screen "Manual.General" 800x480, template "TemplateWithClockAndBackBtnForManual"
   on GenerateScreen: SetBit("Maintenance")
   on ClearScreen: ResetBit("Maintenance")
   GraphicIOField "PlotLight_Round_G" at 224,264 size 24x24; PictureOff "PilotLight_Round_G_Off_256c"; PictureOn "PilotLight_Round_G_On_256c"
      ProcessValue <- "Prezenta aer"
   TextField "Text field_1" at 8,266 size 90x20; Text 'Prezenta aer'
   GraphicIOField "PlotLight_Round_G_1" at 224,48 size 24x24; PictureOn "PilotLight_Round_G_On_256c"; PictureOff "PilotLight_Round_G_Off_256c"
      ProcessValue <- "Aliniere palet"
   TextField "Text field_2" at 8,50 size 91x20; Text 'Aliniere palet'
   GraphicIOField "PlotLight_Round_G_2" at 224,72 size 24x24; PictureOff "PilotLight_Round_G_Off_256c"; PictureOn "PilotLight_Round_G_On_256c"
      ProcessValue <- "Centror extins"
   TextField "Text field_3" at 8,74 size 98x20; Text 'Centror extins'
   GraphicIOField "PlotLight_Round_G_3" at 224,96 size 24x24; PictureOff "PilotLight_Round_G_Off_256c"; PictureOn "PilotLight_Round_G_On_256c"
      ProcessValue <- "Centror retras"
   TextField "Text field_4" at 8,98 size 100x20; Text 'Centror retras'
   GraphicIOField "PlotLight_Round_G_4" at 224,120 size 24x24; PictureOff "PilotLight_Round_G_Off_256c"; PictureOn "PilotLight_Round_G_On_256c"
      ProcessValue <- "Detectie 1 aliniament palet"
   TextField "Text field_5" at 8,122 size 179x20; Text 'Detectie 1 aliniament palet'
   GraphicIOField "PlotLight_Round_G_5" at 224,144 size 24x24; PictureOff "PilotLight_Round_G_Off_256c"; PictureOn "PilotLight_Round_G_On_256c"
      ProcessValue <- "Detectie 2 aliniament palet"
   TextField "Text field_6" at 8,146 size 179x20; Text 'Detectie 2 aliniament palet'
   GraphicIOField "PlotLight_Round_G_6" at 224,168 size 24x24; PictureOff "PilotLight_Round_G_Off_256c"; PictureOn "PilotLight_Round_G_On_256c"
      ProcessValue <- "Detectie palet"
   TextField "Text field_7" at 8,170 size 97x20; Text 'Detectie palet'
   GraphicIOField "PlotLight_Round_G_7" at 224,192 size 24x24; PictureOn "PilotLight_Round_G_On_256c"; PictureOff "PilotLight_Round_G_Off_256c"
      ProcessValue <- "Feed palet"
   TextField "Text field_8" at 8,194 size 72x20; Text 'Feed palet'
   GraphicIOField "PlotLight_Round_G_8" at 224,216 size 24x24; PictureOn "PilotLight_Round_G_On_256c"; PictureOff "PilotLight_Round_G_Off_256c"
      ProcessValue <- "Inaltime maxima"
   TextField "Text field_9" at 8,218 size 109x20; Text 'Inaltime maxima'
   GraphicIOField "PlotLight_Round_G_9" at 224,240 size 24x24; PictureOn "PilotLight_Round_G_On_256c"; PictureOff "PilotLight_Round_G_Off_256c"
      ProcessValue <- "Masurare lungime"
   TextField "Text field_10" at 8,242 size 120x20; Text 'Masurare lungime'
   GraphicIOField "PlotLight_Round_G_10" at 224,288 size 24x24; PictureOn "PilotLight_Round_G_On_256c"; PictureOff "PilotLight_Round_G_Off_256c"
      ProcessValue <- "Prezenta palet iesire"
   TextField "Text field_11" at 8,290 size 140x20; Text 'Prezenta palet iesire'
   GraphicIOField "PlotLight_Round_G_11" at 224,312 size 24x24; PictureOn "PilotLight_Round_G_On_256c"; PictureOff "PilotLight_Round_G_Off_256c"
      ProcessValue <- "Prezenta palet_capat_conveyor"
   TextField "Text field_12" at 8,314 size 215x20; Text 'Prezenta palet_capat_conveyor'
   GraphicIOField "PlotLight_Round_G_12" at 224,336 size 24x24; PictureOn "PilotLight_Round_G_On_256c"; PictureOff "PilotLight_Round_G_Off_256c"
      ProcessValue <- "Prezenta palet_centror"
   TextField "Text field_13" at 8,338 size 158x20; Text 'Prezenta palet_centror'
   GraphicIOField "PlotLight_Round_G_13" at 224,360 size 24x24; PictureOn "PilotLight_Round_G_On_256c"; PictureOff "PilotLight_Round_G_Off_256c"
      ProcessValue <- "Prezenta palet_dreapta"
   TextField "Text field_14" at 8,362 size 161x20; Text 'Prezenta palet_dreapta'
   GraphicIOField "PlotLight_Round_G_14" at 504,264 size 24x24; PictureOn "PilotLight_Round_G_On_256c"; PictureOff "PilotLight_Round_G_Off_256c"
      ProcessValue <- "Protectie cuplata Post reparatii minore"
   TextField "Text field_15" at 264,266 size 230x20; Text 'Prot. cuplata Post reparatii minore'
   GraphicIOField "PlotLight_Round_G_15" at 504,48 size 24x24; PictureOff "PilotLight_Round_G_Off_256c"; PictureOn "PilotLight_Round_G_On_256c"
      ProcessValue <- "Prezenta palet_stanga"
   TextField "Text field_16" at 264,50 size 154x20; Text 'Prezenta palet_stanga'
   GraphicIOField "PlotLight_Round_G_16" at 504,72 size 24x24; PictureOn "PilotLight_Round_G_On_256c"; PictureOff "PilotLight_Round_G_Off_256c"
      ProcessValue <- "Prezenta stiva"
   TextField "Text field_17" at 264,74 size 100x20; Text 'Prezenta stiva'
   GraphicIOField "PlotLight_Round_G_17" at 504,96 size 24x24; PictureOn "PilotLight_Round_G_On_256c"; PictureOff "PilotLight_Round_G_Off_256c"
      ProcessValue <- "Prezenta_stiva"
   TextField "Text field_18" at 264,98 size 104x20; Text 'Prezenta_stiva'
   GraphicIOField "PlotLight_Round_G_18" at 504,120 size 24x24; PictureOn "PilotLight_Round_G_On_256c"; PictureOff "PilotLight_Round_G_Off_256c"
      ProcessValue <- "Protectie cuplata Circular masa fixa"
   TextField "Text field_19" at 264,122 size 235x20; Text 'Protectie cuplata Circular masa fixa'
   GraphicIOField "PlotLight_Round_G_19" at 504,144 size 24x24; PictureOn "PilotLight_Round_G_On_256c"; PictureOff "PilotLight_Round_G_Off_256c"
      ProcessValue <- "Protectie cuplata HMI"
   TextField "Text field_20" at 264,146 size 146x20; Text 'Protectie cuplata HMI'
   GraphicIOField "PlotLight_Round_G_20" at 504,168 size 24x24; PictureOn "PilotLight_Round_G_On_256c"; PictureOff "PilotLight_Round_G_Off_256c"
      ProcessValue <- "Protectie cuplata Iluminat"
   TextField "Text field_21" at 264,170 size 173x20; Text 'Protectie cuplata Iluminat'
   GraphicIOField "PlotLight_Round_G_21" at 504,192 size 24x24; PictureOff "PilotLight_Round_G_Off_256c"; PictureOn "PilotLight_Round_G_On_256c"
      ProcessValue <- "Protectie cuplata Masina demontare paleti dreapta"
   TextField "Text field_22" at 264,194 size 241x20; Text 'Prot. cuplata Mas. dem. pal. dreapta'
   GraphicIOField "PlotLight_Round_G_22" at 504,216 size 24x24; PictureOff "PilotLight_Round_G_Off_256c"; PictureOn "PilotLight_Round_G_On_256c"
      ProcessValue <- "Protectie cuplata Masina demontare paleti stanga"
   TextField "Text field_23" at 264,218 size 234x20; Text 'Prot. cuplata Mas. dem. pal. stanga'
   GraphicIOField "PlotLight_Round_G_23" at 504,240 size 24x24; PictureOff "PilotLight_Round_G_Off_256c"; PictureOn "PilotLight_Round_G_On_256c"
      ProcessValue <- "Protectie cuplata Post reparatie stanga+dreapta"
   TextField "Text field_24" at 264,242 size 218x20; Text 'Prot. cuplata Post rep. stg.+drp.'
   GraphicIOField "PlotLight_Round_G_24" at 504,288 size 24x24; PictureOff "PilotLight_Round_G_Off_256c"; PictureOn "PilotLight_Round_G_On_256c"
      ProcessValue <- "Protectie cuplata TELE"
   TextField "Text field_25" at 264,290 size 149x20; Text 'Protectie cuplata TELE'
   GraphicIOField "PlotLight_Round_G_25" at 504,312 size 24x24; PictureOff "PilotLight_Round_G_Off_256c"; PictureOn "PilotLight_Round_G_On_256c"
      ProcessValue <- "Prezenta palet_capat_conveyor"
   TextField "Text field_26" at 264,314 size 215x20; Text 'Prezenta palet_capat_conveyor'
   GraphicIOField "PlotLight_Round_G_26" at 504,336 size 24x24; PictureOff "PilotLight_Round_G_Off_256c"; PictureOn "PilotLight_Round_G_On_256c"
      ProcessValue <- "Prezenta palet_centror"
   TextField "Text field_27" at 264,338 size 158x20; Text 'Prezenta palet_centror'
   GraphicIOField "PlotLight_Round_G_27" at 504,360 size 24x24; PictureOff "PilotLight_Round_G_Off_256c"; PictureOn "PilotLight_Round_G_On_256c"
      ProcessValue <- "Prezenta palet_dreapta"
   TextField "Text field_28" at 264,362 size 161x20; Text 'Prezenta palet_dreapta'
   GraphicIOField "PlotLight_Round_G_28" at 760,48 size 24x24; PictureOn "PilotLight_Round_G_On_256c"; PictureOff "PilotLight_Round_G_Off_256c"
      ProcessValue <- "Senzor 1 prezenta stiva"
   TextField "Text field_29" at 544,50 size 161x20; Text 'Senzor 1 prezenta stiva'
   GraphicIOField "PlotLight_Round_G_31" at 760,72 size 24x24; PictureOff "PilotLight_Round_G_Off_256c"; PictureOn "PilotLight_Round_G_On_256c"
      ProcessValue <- "Senzor 1 proximitate softstarter aer zona 2"
   TextField "Text field_32" at 544,74 size 206x20; Text 'Senzor 1 prox. soft. aer zona 2'
   GraphicIOField "PlotLight_Round_G_32" at 760,96 size 24x24; PictureOff "PilotLight_Round_G_Off_256c"; PictureOn "PilotLight_Round_G_On_256c"
      ProcessValue <- "Senzor 2 prezenta stiva"
   TextField "Text field_33" at 544,98 size 161x20; Text 'Senzor 2 prezenta stiva'
   GraphicIOField "PlotLight_Round_G_35" at 760,120 size 24x24; PictureOff "PilotLight_Round_G_Off_256c"; PictureOn "PilotLight_Round_G_On_256c"
      ProcessValue <- "Senzor 2 proximitate softstarter aer zona 2"
   TextField "Text field_36" at 544,122 size 206x20; Text 'Senzor 2 prox. soft. aer zona 2'
   GraphicIOField "PlotLight_Round_G_36" at 760,144 size 24x24; PictureOff "PilotLight_Round_G_Off_256c"; PictureOn "PilotLight_Round_G_On_256c"
      ProcessValue <- "Senzor destacking"
   TextField "Text field_37" at 544,146 size 124x20; Text 'Senzor destacking'
   GraphicIOField "PlotLight_Round_G_37" at 760,168 size 24x24; PictureOn "PilotLight_Round_G_On_256c"; PictureOff "PilotLight_Round_G_Off_256c"
      ProcessValue <- "Senzor stacking"
   TextField "Text field_38" at 544,170 size 108x20; Text 'Senzor stacking'
   GraphicIOField "PlotLight_Round_G_38" at 760,192 size 24x24; PictureOn "PilotLight_Round_G_On_256c"; PictureOff "PilotLight_Round_G_Off_256c"
      ProcessValue <- "Start masurare lungime"
   TextField "Text field_39" at 544,194 size 158x20; Text 'Start masurare lungime'

screen "Manual.StackerConveyors" 800x480, template "TemplateWithClockAndBackBtnForManual"
   on GenerateScreen: SetBit("Maintenance")
   on ClearScreen: ResetBit("Maintenance")
   TextField "Text field_15" at 368,54 size 300x20; Text 'Cuplare contactor VFD Conveior 4 descarcare'
   TextField "Text field_16" at 368,94 size 297x20; Text 'Fault Aknowledge VFD Conveior 4 descarcare'
   TextField "Text field_17" at 368,134 size 237x20; Text 'ON/OFF1 VFD Conveior 4 descarcare'
   Switch "Switch_1" at 696,48 size 64x32; CaptionText 'Switch'; TextOff 'OFF'; TextOn 'ON'
      ProcessValue <- "Cuplare contactor VFD Conveior 4 descarcare stacker"
      on SwitchOn: SetBit("Cuplare contactor VFD Conveior 4 descarcare stacker")
      on SwitchOff: ResetBit("Cuplare contactor VFD Conveior 4 descarcare stacker")
   GraphicIOField "PlotLight_Round_G_2" at 288,48 size 24x24; PictureOn "PilotLight_Round_G_On_256c"; PictureOff "PilotLight_Round_G_Off_256c"
      ProcessValue <- "Avarie Conveior 4 stacker"
   TextField "Text field_3" at 16,50 size 174x20; Text 'Avarie Conveior 4 stacker'
   GraphicIOField "PlotLight_Round_G_4" at 288,72 size 24x24; PictureOn "PilotLight_Round_G_On_256c"; PictureOff "PilotLight_Round_G_Off_256c"
      ProcessValue <- "Contactor cuplat Conveior 4 descarcare stacker"
   TextField "Text field_5" at 16,74 size 264x20; Text 'Contactor cuplat Conveior 4 descarcare'
   GraphicIOField "PlotLight_Round_G_6" at 288,120 size 24x24; PictureOn "PilotLight_Round_G_On_256c"; PictureOff "PilotLight_Round_G_Off_256c"
      ProcessValue <- "Frana decuplata Conveior 4 descarcare stacker"
   TextField "Text field_7" at 16,122 size 259x20; Text 'Frana decuplata Conveior 4 descarcare'
   GraphicIOField "PlotLight_Round_G_8" at 288,96 size 24x24; PictureOn "PilotLight_Round_G_On_256c"; PictureOff "PilotLight_Round_G_Off_256c"
      ProcessValue <- "Emergency Stop Stacker"
   TextField "Text field_9" at 16,98 size 164x20; Text 'Emergency Stop Stacker'
   GraphicIOField "PlotLight_Round_G_11" at 288,144 size 24x24; PictureOn "PilotLight_Round_G_On_256c"; PictureOff "PilotLight_Round_G_Off_256c"
      ProcessValue <- "Functionare Conveior 4 stacker"
   TextField "Text field_12" at 16,146 size 207x20; Text 'Functionare Conveior 4 stacker'
   Switch "Switch_3" at 696,88 size 64x32; CaptionText 'Switch'; TextOff 'OFF'; TextOn 'ON'
      ProcessValue <- "Fault Aknowledge VFD Conveior 4 descarcare stacker"
      on SwitchOn: SetBit("Fault Aknowledge VFD Conveior 4 descarcare stacker")
      on SwitchOff: ResetBit("Fault Aknowledge VFD Conveior 4 descarcare stacker")
   Switch "Switch_4" at 696,128 size 64x32; CaptionText 'Switch'; TextOff 'OFF'; TextOn 'ON'
      ProcessValue <- "ON/OFF1 VFD Conveior 4 descarcare stacker"
      on SwitchOn: SetBit("ON/OFF1 VFD Conveior 4 descarcare stacker")
      on SwitchOff: ResetBit("ON/OFF1 VFD Conveior 4 descarcare stacker")
   GraphicIOField "PlotLight_Round_G_1" at 288,168 size 24x24; PictureOff "PilotLight_Round_G_Off_256c"; PictureOn "PilotLight_Round_G_On_256c"
      ProcessValue <- "Protectie cuplata Conveior 4 descarcare stacker"
   TextField "Text field_1" at 16,170 size 267x20; Text 'Protectie cuplata Conveior 4 descarcare'

screen "Manual.Safety" 800x480, template "TemplateWithClockAndBackBtnForManual"
   on GenerateScreen: SetBit("Maintenance")
   on ClearScreen: ResetBit("Maintenance")
   GraphicIOField "PlotLight_Round_G_2" at 280,48 size 24x24; PictureOn "PilotLight_Round_G_On_256c"; PictureOff "PilotLight_Round_G_Off_256c"
      ProcessValue <- "Destacker 110KF1 Safety Relay"
   TextField "Text field_3" at 16,50 size 208x20; Text 'Destacker 110KF1 Safety Relay'
   GraphicIOField "PlotLight_Round_G_1" at 280,72 size 24x24; PictureOff "PilotLight_Round_G_Off_256c"; PictureOn "PilotLight_Round_G_On_256c"
      ProcessValue <- "Destacker 111KF1 Safety Barrier Relay"
   TextField "Text field_1" at 16,74 size 257x20; Text 'Destacker 111KF1 Safety Barrier Relay'
   GraphicIOField "PlotLight_Round_G_3" at 280,96 size 24x24; PictureOn "PilotLight_Round_G_On_256c"; PictureOff "PilotLight_Round_G_Off_256c"
      ProcessValue <- "Emergency Stop Destacker"
   TextField "Text field_2" at 16,98 size 180x20; Text 'Emergency Stop Destacker'
   GraphicIOField "PlotLight_Round_G_4" at 280,120 size 24x24; PictureOff "PilotLight_Round_G_Off_256c"; PictureOn "PilotLight_Round_G_On_256c"
      ProcessValue <- "Emergency Stop Stacker"
   TextField "Text field_4" at 16,122 size 164x20; Text 'Emergency Stop Stacker'
   GraphicIOField "PlotLight_Round_G_5" at 280,144 size 24x24; PictureOff "PilotLight_Round_G_Off_256c"; PictureOn "PilotLight_Round_G_On_256c"
      ProcessValue <- "Emergency Stop Zone 2"
   TextField "Text field_5" at 16,146 size 157x20; Text 'Emergency Stop Zone 2'
   GraphicIOField "PlotLight_Round_G_6" at 280,168 size 24x24; PictureOff "PilotLight_Round_G_Off_256c"; PictureOn "PilotLight_Round_G_On_256c"
      ProcessValue <- "Stacker 113KF1 Safety Relay"
   TextField "Text field_6" at 16,170 size 192x20; Text 'Stacker 113KF1 Safety Relay'
   GraphicIOField "PlotLight_Round_G_7" at 280,192 size 24x24; PictureOff "PilotLight_Round_G_Off_256c"; PictureOn "PilotLight_Round_G_On_256c"
      ProcessValue <- "Stacker 114KF1 Safety Barrier Relay 1"
   TextField "Text field_7" at 16,194 size 253x20; Text 'Stacker 114KF1 Safety Barrier Relay 1'
   GraphicIOField "PlotLight_Round_G_8" at 280,216 size 24x24; PictureOff "PilotLight_Round_G_Off_256c"; PictureOn "PilotLight_Round_G_On_256c"
      ProcessValue <- "Stacker 115KF1 Safety Barrier Relay 2"
   TextField "Text field_8" at 16,218 size 253x20; Text 'Stacker 115KF1 Safety Barrier Relay 2'
   GraphicIOField "PlotLight_Round_G_9" at 280,240 size 24x24; PictureOff "PilotLight_Round_G_Off_256c"; PictureOn "PilotLight_Round_G_On_256c"
      ProcessValue <- "Zone 2 112KF1 Safety Relay"
   TextField "Text field_9" at 16,242 size 185x20; Text 'Zone 2 112KF1 Safety Relay'
   TextField "Text field_14" at 384,54 size 250x20; Text 'Reset Destacker 110KF1 Safety Relay'
   Switch "Switch_2" at 696,48 size 64x32; CaptionText 'Switch'; TextOff 'OFF'; TextOn 'ON'
      ProcessValue <- "Reset Destacker 110KF1 Safety Relay"
      on SwitchOn: SetBit("Reset Destacker 110KF1 Safety Relay")
      on SwitchOff: ResetBit("Reset Destacker 110KF1 Safety Relay")
   TextField "Text field_10" at 384,94 size 299x20; Text 'Reset Destacker 111KF1 Safety Barrier Relay'
   Switch "Switch_1" at 696,88 size 64x32; CaptionText 'Switch'; TextOff 'OFF'; TextOn 'ON'
      ProcessValue <- "Reset Destacker 111KF1 Safety Barrier Relay"
      on SwitchOn: SetBit("Reset Destacker 111KF1 Safety Barrier Relay")
      on SwitchOff: ResetBit("Reset Destacker 111KF1 Safety Barrier Relay")
   TextField "Text field_11" at 384,134 size 136x20; Text 'Reset safety Zone 2'
   Switch "Switch_3" at 696,128 size 64x32; CaptionText 'Switch'; TextOff 'OFF'; TextOn 'ON'
      ProcessValue <- "Reset safety Zone 2"
      on SwitchOn: SetBit("Reset safety Zone 2")
      on SwitchOff: ResetBit("Reset safety Zone 2")
   TextField "Text field_12" at 384,174 size 234x20; Text 'Reset Stacker 113KF1 Safety Relay'
   Switch "Switch_4" at 696,168 size 64x32; CaptionText 'Switch'; TextOff 'OFF'; TextOn 'ON'
      ProcessValue <- "Reset Stacker 113KF1 Safety Relay"
      on SwitchOn: SetBit("Reset Stacker 113KF1 Safety Relay")
      on SwitchOff: ResetBit("Reset Stacker 113KF1 Safety Relay")
   TextField "Text field_13" at 384,214 size 295x20; Text 'Reset Stacker 114KF1 Safety Barrier Relay 1'
   Switch "Switch_5" at 696,208 size 64x32; CaptionText 'Switch'; TextOff 'OFF'; TextOn 'ON'
      ProcessValue <- "Reset Stacker 114KF1 Safety Barrier Relay 1"
      on SwitchOn: SetBit("Reset Stacker 114KF1 Safety Barrier Relay 1")
      on SwitchOff: ResetBit("Reset Stacker 114KF1 Safety Barrier Relay 1")
   TextField "Text field_15" at 384,254 size 295x20; Text 'Reset Stacker 115KF1 Safety Barrier Relay 2'
   Switch "Switch_6" at 696,248 size 64x32; CaptionText 'Switch'; TextOff 'OFF'; TextOn 'ON'
      ProcessValue <- "Reset Stacker 115KF1 Safety Barrier Relay 2"
      on SwitchOn: SetBit("Reset Stacker 115KF1 Safety Barrier Relay 2")
      on SwitchOff: ResetBit("Reset Stacker 115KF1 Safety Barrier Relay 2")
   TextField "Text field_16" at 384,294 size 227x20; Text 'Reset Zone 2 112KF1 Safety Relay'
   Switch "Switch_7" at 696,288 size 64x32; CaptionText 'Switch'; TextOff 'OFF'; TextOn 'ON'
      ProcessValue <- "Reset Zone 2 112KF1 Safety Relay"
      on SwitchOn: SetBit("Reset Zone 2 112KF1 Safety Relay")
      on SwitchOff: ResetBit("Reset Zone 2 112KF1 Safety Relay")

screen "Manual.DestackerConveyors" 800x480, template "TemplateWithClockAndBackBtnForManual"
   on GenerateScreen: SetBit("Maintenance")
   on ClearScreen: ResetBit("Maintenance")
   TextField "Text field_15" at 368,54 size 296x20; Text 'Cuplare contactor VFD Conveior 1 alimentare'
   TextField "Text field_16" at 368,94 size 293x20; Text 'Fault Aknowledge VFD Conveior 1 alimentare'
   TextField "Text field_17" at 368,134 size 233x20; Text 'ON/OFF1 VFD Conveior 1 alimentare'
   TextField "Text field_18" at 368,174 size 262x20; Text 'Cuplare contactor VFD Conveior 2 iesire'
   TextField "Text field_19" at 368,214 size 259x20; Text 'Fault Aknowledge VFD Conveior 2 iesire'
   TextField "Text field_20" at 368,254 size 199x20; Text 'ON/OFF1 VFD Conveior 2 iesire'
   Switch "Switch_1" at 696,48 size 64x32; CaptionText 'Switch'; TextOff 'OFF'; TextOn 'ON'
      ProcessValue <- "Cuplare contactor VFD Conveior 1 alimentare destacker"
      on SwitchOn: SetBit("Cuplare contactor VFD Conveior 1 alimentare destacker")
      on SwitchOff: ResetBit("Cuplare contactor VFD Conveior 1 alimentare destacker")
   GraphicIOField "PlotLight_Round_G" at 280,144 size 24x24; PictureOff "PilotLight_Round_G_Off_256c"; PictureOn "PilotLight_Round_G_On_256c"
      ProcessValue <- "Protectie cuplata Conveior 1 alimentare destacker"
   TextField "Text field_1" at 16,146 size 263x20; Text 'Protectie cuplata Conveior 1 alimentare'
   GraphicIOField "PlotLight_Round_G_1" at 280,264 size 24x24; PictureOn "PilotLight_Round_G_On_256c"; PictureOff "PilotLight_Round_G_Off_256c"
      ProcessValue <- "Protectie cuplata Conveior 2 iesire destacker"
   TextField "Text field_2" at 16,266 size 229x20; Text 'Protectie cuplata Conveior 2 iesire'
   GraphicIOField "PlotLight_Round_G_2" at 280,48 size 24x24; PictureOff "PilotLight_Round_G_Off_256c"; PictureOn "PilotLight_Round_G_On_256c"
      ProcessValue <- "Avarie Conveior 1 alimentare destacker"
   TextField "Text field_3" at 16,50 size 194x20; Text 'Avarie Conveior 1 alimentare'
   GraphicIOField "PlotLight_Round_G_3" at 280,168 size 24x24; PictureOff "PilotLight_Round_G_Off_256c"; PictureOn "PilotLight_Round_G_On_256c"
      ProcessValue <- "Avarie Conveior 2 iesire destacker"
   TextField "Text field_4" at 16,170 size 160x20; Text 'Avarie Conveior 2 iesire'
   GraphicIOField "PlotLight_Round_G_4" at 280,72 size 24x24; PictureOff "PilotLight_Round_G_Off_256c"; PictureOn "PilotLight_Round_G_On_256c"
      ProcessValue <- "Contactor cuplat Conveior 1 alimentare destacker"
   TextField "Text field_5" at 16,74 size 260x20; Text 'Contactor cuplat Conveior 1 alimentare'
   GraphicIOField "PlotLight_Round_G_5" at 280,192 size 24x24; PictureOff "PilotLight_Round_G_Off_256c"; PictureOn "PilotLight_Round_G_On_256c"
      ProcessValue <- "Contactor cuplat Conveior 2 iesire destacker"
   TextField "Text field_6" at 16,194 size 226x20; Text 'Contactor cuplat Conveior 2 iesire'
   GraphicIOField "PlotLight_Round_G_6" at 280,96 size 24x24; PictureOff "PilotLight_Round_G_Off_256c"; PictureOn "PilotLight_Round_G_On_256c"
      ProcessValue <- "Frana decuplata Conveior 1 alimentare destacker"
   TextField "Text field_7" at 16,98 size 255x20; Text 'Frana decuplata Conveior 1 alimentare'
   GraphicIOField "PlotLight_Round_G_7" at 280,216 size 24x24; PictureOff "PilotLight_Round_G_Off_256c"; PictureOn "PilotLight_Round_G_On_256c"
      ProcessValue <- "Frana decuplata Conveior 2 iesire destacker"
   TextField "Text field_8" at 16,218 size 221x20; Text 'Frana decuplata Conveior 2 iesire'
   GraphicIOField "PlotLight_Round_G_8" at 280,120 size 24x24; PictureOff "PilotLight_Round_G_Off_256c"; PictureOn "PilotLight_Round_G_On_256c"
      ProcessValue <- "Functionare Conveior 1 alimentare destacker"
   TextField "Text field_9" at 16,122 size 227x20; Text 'Functionare Conveior 1 alimentare'
   GraphicIOField "PlotLight_Round_G_9" at 280,240 size 24x24; PictureOff "PilotLight_Round_G_Off_256c"; PictureOn "PilotLight_Round_G_On_256c"
      ProcessValue <- "Functionare Conveior 2 iesire destacker"
   TextField "Text field_10" at 16,242 size 193x20; Text 'Functionare Conveior 2 iesire'
   GraphicIOField "PlotLight_Round_G_10" at 280,288 size 24x24; PictureOff "PilotLight_Round_G_Off_256c"; PictureOn "PilotLight_Round_G_On_256c"
      ProcessValue <- "Senzor 1 proximitate softstarter aer destacker"
   TextField "Text field_11" at 16,290 size 243x20; Text 'Senzor 1 proximitate softstarter aer'
   GraphicIOField "PlotLight_Round_G_11" at 280,336 size 24x24; PictureOff "PilotLight_Round_G_Off_256c"; PictureOn "PilotLight_Round_G_On_256c"
      ProcessValue <- "Reset safety Destacker"
   TextField "Text field_12" at 16,338 size 89x20; Text 'Reset safety'
   GraphicIOField "PlotLight_Round_G_12" at 280,312 size 24x24; PictureOff "PilotLight_Round_G_Off_256c"; PictureOn "PilotLight_Round_G_On_256c"
      ProcessValue <- "Senzor 2 proximitate softstarter aer destacker"
   TextField "Text field_13" at 16,314 size 243x20; Text 'Senzor 2 proximitate softstarter aer'
   Switch "Switch_3" at 696,88 size 64x32; CaptionText 'Switch'; TextOff 'OFF'; TextOn 'ON'
      ProcessValue <- "Fault Aknowledge VFD Conveior 1 alimentare destacker"
      on SwitchOn: SetBit("Fault Aknowledge VFD Conveior 1 alimentare destacker")
      on SwitchOff: ResetBit("Fault Aknowledge VFD Conveior 1 alimentare destacker")
   Switch "Switch_4" at 696,128 size 64x32; CaptionText 'Switch'; TextOff 'OFF'; TextOn 'ON'
      ProcessValue <- "ON/OFF1 VFD Conveior 1 alimentare destacker"
      on SwitchOn: SetBit("ON/OFF1 VFD Conveior 1 alimentare destacker")
      on SwitchOff: ResetBit("ON/OFF1 VFD Conveior 1 alimentare destacker")
   Switch "Switch_5" at 696,168 size 64x32; CaptionText 'Switch'; TextOff 'OFF'; TextOn 'ON'
      ProcessValue <- "Cuplare contactor VFD Conveior 2 iesire destacker"
      on SwitchOn: SetBit("Cuplare contactor VFD Conveior 2 iesire destacker")
      on SwitchOff: ResetBit("Cuplare contactor VFD Conveior 2 iesire destacker")
   Switch "Switch_6" at 696,208 size 64x32; CaptionText 'Switch'; TextOff 'OFF'; TextOn 'ON'
      ProcessValue <- "Fault Aknowledge VFD Conveior 2 iesire destacker"
      on SwitchOn: SetBit("Fault Aknowledge VFD Conveior 2 iesire destacker")
      on SwitchOff: ResetBit("Fault Aknowledge VFD Conveior 2 iesire destacker")
   Switch "Switch_7" at 696,248 size 64x32; CaptionText 'Switch'; TextOff 'OFF'; TextOn 'ON'
      ProcessValue <- "ON/OFF1 VFD Conveior 2 iesire destacker"
      on SwitchOn: SetBit("ON/OFF1 VFD Conveior 2 iesire destacker")
      on SwitchOff: ResetBit("ON/OFF1 VFD Conveior 2 iesire destacker")

screen "Manual.Transfer" 800x480, template "TemplateWithClockAndBackBtnForManual"
   on GenerateScreen: SetBit("Maintenance")
   on ClearScreen: ResetBit("Maintenance")
   TextField "Text field_14" at 368,54 size 330x20; Text 'Cuplare contactor VFD Conveior 3 transfer palet 2'
   TextField "Text field_15" at 368,94 size 327x20; Text 'Fault Aknowledge VFD Conveior 3 transfer palet 2'
   TextField "Text field_16" at 368,134 size 289x20; Text 'Frana decuplata Conveior 3 transfer palet 2'
   TextField "Text field_17" at 368,174 size 267x20; Text 'ON/OFF1 VFD Conveior 3 transfer palet 2'
   TextField "Text field_18" at 368,214 size 322x20; Text 'Softstarter aer 1.1 Conveior 1 preluare paleti OK'
   TextField "Text field_19" at 368,254 size 322x20; Text 'Softstarter aer 1.2 Conveior 1 preluare paleti OK'
   TextField "Text field_20" at 368,294 size 232x20; Text 'Start Conveior 1 preluare paleti OK'
   Switch "Switch_1" at 696,88 size 64x32; CaptionText 'Switch'; TextOff 'OFF'; TextOn 'ON'
      ProcessValue <- "Fault Aknowledge VFD Conveior 3 transfer palet 2"
      on SwitchOn: SetBit("Fault Aknowledge VFD Conveior 3 transfer palet 2")
      on SwitchOff: ResetBit("Fault Aknowledge VFD Conveior 3 transfer palet 2")
   GraphicIOField "PlotLight_Round_G" at 328,144 size 24x24; PictureOn "PilotLight_Round_G_On_256c"; PictureOff "PilotLight_Round_G_Off_256c"
      ProcessValue <- "Functionare Conveior 2 transfer palet 1"
   TextField "Text field_1" at 16,146 size 261x20; Text 'Functionare Conveior 2 transfer palet 1'
   GraphicIOField "PlotLight_Round_G_2" at 328,48 size 24x24; PictureOn "PilotLight_Round_G_On_256c"; PictureOff "PilotLight_Round_G_Off_256c"
      ProcessValue <- "Avarie Conveior 3 transfer palet 2"
   TextField "Text field_3" at 16,50 size 228x20; Text 'Avarie Conveior 3 transfer palet 2'
   GraphicIOField "PlotLight_Round_G_3" at 328,168 size 24x24; PictureOn "PilotLight_Round_G_On_256c"; PictureOff "PilotLight_Round_G_Off_256c"
      ProcessValue <- "Functionare Conveior 3 transfer palet 2"
   TextField "Text field_4" at 16,170 size 261x20; Text 'Functionare Conveior 3 transfer palet 2'
   GraphicIOField "PlotLight_Round_G_4" at 328,72 size 24x24; PictureOn "PilotLight_Round_G_On_256c"; PictureOff "PilotLight_Round_G_Off_256c"
      ProcessValue <- "Contactor cuplat Conveior 3 transfer palet 2"
   TextField "Text field_5" at 16,74 size 294x20; Text 'Contactor cuplat Conveior 3 transfer palet 2'
   GraphicIOField "PlotLight_Round_G_5" at 328,192 size 24x24; PictureOn "PilotLight_Round_G_On_256c"; PictureOff "PilotLight_Round_G_Off_256c"
      ProcessValue <- "Protectie cuplata Conveior 1 preluare paleti OK"
   TextField "Text field_6" at 16,194 size 310x20; Text 'Protectie cuplata Conveior 1 preluare paleti OK'
   GraphicIOField "PlotLight_Round_G_6" at 328,96 size 24x24; PictureOn "PilotLight_Round_G_On_256c"; PictureOff "PilotLight_Round_G_Off_256c"
      ProcessValue <- "Frana decuplata Conveior 3 transfer palet 2"
   TextField "Text field_7" at 16,98 size 289x20; Text 'Frana decuplata Conveior 3 transfer palet 2'
   GraphicIOField "PlotLight_Round_G_7" at 328,216 size 24x24; PictureOn "PilotLight_Round_G_On_256c"; PictureOff "PilotLight_Round_G_Off_256c"
      ProcessValue <- "Protectie cuplata Conveior 2 transfer palet 1"
   TextField "Text field_8" at 16,218 size 297x20; Text 'Protectie cuplata Conveior 2 transfer palet 1'
   GraphicIOField "PlotLight_Round_G_8" at 328,120 size 24x24; PictureOn "PilotLight_Round_G_On_256c"; PictureOff "PilotLight_Round_G_Off_256c"
      ProcessValue <- "Functionare Conveior 1 preluare paleti OK"
   TextField "Text field_9" at 16,122 size 274x20; Text 'Functionare Conveior 1 preluare paleti OK'
   GraphicIOField "PlotLight_Round_G_9" at 328,240 size 24x24; PictureOn "PilotLight_Round_G_On_256c"; PictureOff "PilotLight_Round_G_Off_256c"
      ProcessValue <- "Protectie cuplata Conveior 3 transfer palet 2"
   TextField "Text field_10" at 16,242 size 297x20; Text 'Protectie cuplata Conveior 3 transfer palet 2'
   Switch "Switch_2" at 696,48 size 64x32; CaptionText 'Switch'; TextOff 'OFF'; TextOn 'ON'
      ProcessValue <- "Cuplare contactor VFD Conveior 3 transfer palet 2"
      on SwitchOn: SetBit("Cuplare contactor VFD Conveior 3 transfer palet 2")
      on SwitchOff: ResetBit("Cuplare contactor VFD Conveior 3 transfer palet 2")
   Switch "Switch_3" at 696,128 size 64x32; CaptionText 'Switch'; TextOff 'OFF'; TextOn 'ON'
      ProcessValue <- "Frana decuplata Conveior 3 transfer palet 2"
   Switch "Switch_4" at 696,168 size 64x32; CaptionText 'Switch'; TextOff 'OFF'; TextOn 'ON'
      ProcessValue <- "ON/OFF1 VFD Conveior 3 transfer palet 2"
      on SwitchOn: SetBit("ON/OFF1 VFD Conveior 3 transfer palet 2")
      on SwitchOff: ResetBit("ON/OFF1 VFD Conveior 3 transfer palet 2")
   Switch "Switch_5" at 696,208 size 64x32; CaptionText 'Switch'; TextOff 'OFF'; TextOn 'ON'
      ProcessValue <- "Softstarter aer 1.1 Conveior 1 preluare paleti OK"
      on SwitchOn: SetBit("Softstarter aer 1.1 Conveior 1 preluare paleti OK")
      on SwitchOff: ResetBit("Softstarter aer 1.1 Conveior 1 preluare paleti OK")
   Switch "Switch_6" at 696,248 size 64x32; CaptionText 'Switch'; TextOff 'OFF'; TextOn 'ON'
      ProcessValue <- "Softstarter aer 1.2 Conveior 1 preluare paleti OK"
      on SwitchOn: SetBit("Softstarter aer 1.2 Conveior 1 preluare paleti OK")
      on SwitchOff: ResetBit("Softstarter aer 1.2 Conveior 1 preluare paleti OK")
   Switch "Switch_7" at 696,288 size 64x32; CaptionText 'Switch'; TextOff 'OFF'; TextOn 'ON'
      on SwitchOn: SetBit("Start Conveior 1 preluare paleti OK")
      on SwitchOff: ResetBit("Start Conveior 1 preluare paleti OK")
   TextField "Text field_2" at 368,334 size 219x20; Text 'Start Conveior 2 transfer palet 1'
   Switch "Switch_8" at 696,328 size 64x32; CaptionText 'Switch'; TextOff 'OFF'; TextOn 'ON'
      ProcessValue <- "Start Conveior 2 transfer palet 1"
      on SwitchOn: SetBit("Start Conveior 2 transfer palet 1")
      on SwitchOff: ResetBit("Start Conveior 2 transfer palet 1")

screen "Manual.IOLinkDiag" 800x480, template "TemplateWithClockAndBackBtnForManual"
   on GenerateScreen: SetBit("Maintenance")
   on ClearScreen: ResetBit("Maintenance")
   GraphicIOField "PlotLight_Round_G" at 136,48 size 24x24; PictureOn "PilotLight_Round_G_On_256c"; PictureOff "PilotLight_Round_G_Off_256c"
      ProcessValue <- "MD_IS1_SC_X1.0"
   TextField "Text field_1" at 8,50 size 115x20; Text 'MD_IS1_SC_X1.0'
   GraphicIOField "PlotLight_Round_G_1" at 136,72 size 24x24; PictureOff "PilotLight_Round_G_Off_256c"; PictureOn "PilotLight_Round_G_On_256c"
      ProcessValue <- "MD_IS1_SC_X1.1"
   TextField "Text field_2" at 8,74 size 115x20; Text 'MD_IS1_SC_X1.1'
   GraphicIOField "PlotLight_Round_G_2" at 136,96 size 24x24; PictureOff "PilotLight_Round_G_Off_256c"; PictureOn "PilotLight_Round_G_On_256c"
      ProcessValue <- "MD_IS1_SC_X1.2"
   TextField "Text field_3" at 8,98 size 115x20; Text 'MD_IS1_SC_X1.2'
   GraphicIOField "PlotLight_Round_G_3" at 136,120 size 24x24; PictureOn "PilotLight_Round_G_On_256c"; PictureOff "PilotLight_Round_G_Off_256c"
      ProcessValue <- "MD_IS1_SC_X1.3"
   TextField "Text field_4" at 8,122 size 115x20; Text 'MD_IS1_SC_X1.3'
   GraphicIOField "PlotLight_Round_G_4" at 136,144 size 24x24; PictureOn "PilotLight_Round_G_On_256c"; PictureOff "PilotLight_Round_G_Off_256c"
      ProcessValue <- "MD_IS1_SC_X1.4"
   TextField "Text field_5" at 8,146 size 115x20; Text 'MD_IS1_SC_X1.4'
   GraphicIOField "PlotLight_Round_G_5" at 136,168 size 24x24; PictureOn "PilotLight_Round_G_On_256c"; PictureOff "PilotLight_Round_G_Off_256c"
      ProcessValue <- "MD_IS1_SC_X1.5"
   TextField "Text field_6" at 8,170 size 115x20; Text 'MD_IS1_SC_X1.5'
   GraphicIOField "PlotLight_Round_G_6" at 136,192 size 24x24; PictureOn "PilotLight_Round_G_On_256c"; PictureOff "PilotLight_Round_G_Off_256c"
      ProcessValue <- "MD_IS1_SC_X1.6"
   TextField "Text field_7" at 8,194 size 115x20; Text 'MD_IS1_SC_X1.6'
   GraphicIOField "PlotLight_Round_G_7" at 136,216 size 24x24; PictureOn "PilotLight_Round_G_On_256c"; PictureOff "PilotLight_Round_G_Off_256c"
      ProcessValue <- "MD_IS1_SC_X1.7"
   TextField "Text field_8" at 8,218 size 115x20; Text 'MD_IS1_SC_X1.7'
   GraphicIOField "PlotLight_Round_G_8" at 312,48 size 24x24; PictureOff "PilotLight_Round_G_Off_256c"; PictureOn "PilotLight_Round_G_On_256c"
      ProcessValue <- "MD_IS2_SC_X1.0"
   TextField "Text field_9" at 184,50 size 115x20; Text 'MD_IS2_SC_X1.0'
   GraphicIOField "PlotLight_Round_G_9" at 312,72 size 24x24; PictureOn "PilotLight_Round_G_On_256c"; PictureOff "PilotLight_Round_G_Off_256c"
      ProcessValue <- "MD_IS2_SC_X1.1"
   TextField "Text field_10" at 184,74 size 115x20; Text 'MD_IS2_SC_X1.1'
   GraphicIOField "PlotLight_Round_G_10" at 312,96 size 24x24; PictureOn "PilotLight_Round_G_On_256c"; PictureOff "PilotLight_Round_G_Off_256c"
      ProcessValue <- "MD_IS2_SC_X1.2"
   TextField "Text field_11" at 184,98 size 115x20; Text 'MD_IS2_SC_X1.2'
   GraphicIOField "PlotLight_Round_G_11" at 312,120 size 24x24; PictureOff "PilotLight_Round_G_Off_256c"; PictureOn "PilotLight_Round_G_On_256c"
      ProcessValue <- "MD_IS2_SC_X1.3"
   TextField "Text field_12" at 184,122 size 115x20; Text 'MD_IS2_SC_X1.3'
   GraphicIOField "PlotLight_Round_G_12" at 312,144 size 24x24; PictureOff "PilotLight_Round_G_Off_256c"; PictureOn "PilotLight_Round_G_On_256c"
      ProcessValue <- "MD_IS2_SC_X1.4"
   TextField "Text field_13" at 184,146 size 115x20; Text 'MD_IS2_SC_X1.4'
   GraphicIOField "PlotLight_Round_G_13" at 312,168 size 24x24; PictureOff "PilotLight_Round_G_Off_256c"; PictureOn "PilotLight_Round_G_On_256c"
      ProcessValue <- "MD_IS2_SC_X1.5"
   TextField "Text field_14" at 184,170 size 115x20; Text 'MD_IS2_SC_X1.5'
   GraphicIOField "PlotLight_Round_G_14" at 312,192 size 24x24; PictureOff "PilotLight_Round_G_Off_256c"; PictureOn "PilotLight_Round_G_On_256c"
      ProcessValue <- "MD_IS2_SC_X1.6"
   TextField "Text field_15" at 184,194 size 115x20; Text 'MD_IS2_SC_X1.6'
   GraphicIOField "PlotLight_Round_G_15" at 312,216 size 24x24; PictureOff "PilotLight_Round_G_Off_256c"; PictureOn "PilotLight_Round_G_On_256c"
      ProcessValue <- "MD_IS2_SC_X1.7"
   TextField "Text field_16" at 184,218 size 115x20; Text 'MD_IS2_SC_X1.7'
   GraphicIOField "PlotLight_Round_G_16" at 136,240 size 24x24; PictureOn "PilotLight_Round_G_On_256c"; PictureOff "PilotLight_Round_G_Off_256c"
      ProcessValue <- "MD_OS_SC_X1.0"
   TextField "Text field_17" at 8,242 size 111x20; Text 'MD_OS_SC_X1.0'
   GraphicIOField "PlotLight_Round_G_17" at 136,264 size 24x24; PictureOff "PilotLight_Round_G_Off_256c"; PictureOn "PilotLight_Round_G_On_256c"
      ProcessValue <- "MD_OS_SC_X1.1"
   TextField "Text field_18" at 8,266 size 111x20; Text 'MD_OS_SC_X1.1'
   GraphicIOField "PlotLight_Round_G_18" at 136,288 size 24x24; PictureOff "PilotLight_Round_G_Off_256c"; PictureOn "PilotLight_Round_G_On_256c"
      ProcessValue <- "MD_OS_SC_X1.2"
   TextField "Text field_19" at 8,290 size 111x20; Text 'MD_OS_SC_X1.2'
   GraphicIOField "PlotLight_Round_G_19" at 136,312 size 24x24; PictureOn "PilotLight_Round_G_On_256c"; PictureOff "PilotLight_Round_G_Off_256c"
      ProcessValue <- "MD_OS_SC_X1.3"
   TextField "Text field_20" at 8,314 size 111x20; Text 'MD_OS_SC_X1.3'
   GraphicIOField "PlotLight_Round_G_20" at 136,336 size 24x24; PictureOn "PilotLight_Round_G_On_256c"; PictureOff "PilotLight_Round_G_Off_256c"
      ProcessValue <- "MD_OS_SC_X1.4"
   TextField "Text field_21" at 8,338 size 111x20; Text 'MD_OS_SC_X1.4'
   GraphicIOField "PlotLight_Round_G_21" at 136,360 size 24x24; PictureOn "PilotLight_Round_G_On_256c"; PictureOff "PilotLight_Round_G_Off_256c"
      ProcessValue <- "MD_OS_SC_X1.5"
   TextField "Text field_22" at 8,362 size 111x20; Text 'MD_OS_SC_X1.5'
   GraphicIOField "PlotLight_Round_G_22" at 488,48 size 24x24; PictureOff "PilotLight_Round_G_Off_256c"; PictureOn "PilotLight_Round_G_On_256c"
      ProcessValue <- "MS_IS1_SC_X1.0"
   TextField "Text field_23" at 360,50 size 114x20; Text 'MS_IS1_SC_X1.0'
   GraphicIOField "PlotLight_Round_G_23" at 488,72 size 24x24; PictureOn "PilotLight_Round_G_On_256c"; PictureOff "PilotLight_Round_G_Off_256c"
      ProcessValue <- "MS_IS1_SC_X1.1"
   TextField "Text field_24" at 360,74 size 114x20; Text 'MS_IS1_SC_X1.1'
   GraphicIOField "PlotLight_Round_G_24" at 488,96 size 24x24; PictureOn "PilotLight_Round_G_On_256c"; PictureOff "PilotLight_Round_G_Off_256c"
      ProcessValue <- "MS_IS1_SC_X1.2"
   TextField "Text field_25" at 360,98 size 114x20; Text 'MS_IS1_SC_X1.2'
   GraphicIOField "PlotLight_Round_G_25" at 488,120 size 24x24; PictureOff "PilotLight_Round_G_Off_256c"; PictureOn "PilotLight_Round_G_On_256c"
      ProcessValue <- "MS_IS1_SC_X1.3"
   TextField "Text field_26" at 360,122 size 114x20; Text 'MS_IS1_SC_X1.3'
   GraphicIOField "PlotLight_Round_G_26" at 488,144 size 24x24; PictureOff "PilotLight_Round_G_Off_256c"; PictureOn "PilotLight_Round_G_On_256c"
      ProcessValue <- "MS_IS1_SC_X1.4"
   TextField "Text field_27" at 360,146 size 114x20; Text 'MS_IS1_SC_X1.4'
   GraphicIOField "PlotLight_Round_G_27" at 488,168 size 24x24; PictureOff "PilotLight_Round_G_Off_256c"; PictureOn "PilotLight_Round_G_On_256c"
      ProcessValue <- "MS_IS1_SC_X1.5"
   TextField "Text field_28" at 360,170 size 114x20; Text 'MS_IS1_SC_X1.5'
   GraphicIOField "PlotLight_Round_G_28" at 488,192 size 24x24; PictureOff "PilotLight_Round_G_Off_256c"; PictureOn "PilotLight_Round_G_On_256c"
      ProcessValue <- "MS_IS1_SC_X1.6"
   TextField "Text field_29" at 360,194 size 114x20; Text 'MS_IS1_SC_X1.6'
   GraphicIOField "PlotLight_Round_G_29" at 488,216 size 24x24; PictureOff "PilotLight_Round_G_Off_256c"; PictureOn "PilotLight_Round_G_On_256c"
      ProcessValue <- "MS_IS1_SC_X1.7"
   TextField "Text field_30" at 360,218 size 114x20; Text 'MS_IS1_SC_X1.7'
   GraphicIOField "PlotLight_Round_G_30" at 664,48 size 24x24; PictureOn "PilotLight_Round_G_On_256c"; PictureOff "PilotLight_Round_G_Off_256c"
      ProcessValue <- "MS_IS2_SC_X1.0"
   TextField "Text field_31" at 536,50 size 114x20; Text 'MS_IS2_SC_X1.0'
   GraphicIOField "PlotLight_Round_G_31" at 664,72 size 24x24; PictureOff "PilotLight_Round_G_Off_256c"; PictureOn "PilotLight_Round_G_On_256c"
      ProcessValue <- "MS_IS2_SC_X1.1"
   TextField "Text field_32" at 536,74 size 114x20; Text 'MS_IS2_SC_X1.1'
   GraphicIOField "PlotLight_Round_G_32" at 664,96 size 24x24; PictureOff "PilotLight_Round_G_Off_256c"; PictureOn "PilotLight_Round_G_On_256c"
      ProcessValue <- "MS_IS2_SC_X1.2"
   TextField "Text field_33" at 536,98 size 114x20; Text 'MS_IS2_SC_X1.2'
   GraphicIOField "PlotLight_Round_G_33" at 664,120 size 24x24; PictureOn "PilotLight_Round_G_On_256c"; PictureOff "PilotLight_Round_G_Off_256c"
      ProcessValue <- "MS_IS2_SC_X1.3"
   TextField "Text field_34" at 536,122 size 114x20; Text 'MS_IS2_SC_X1.3'
   GraphicIOField "PlotLight_Round_G_34" at 664,144 size 24x24; PictureOn "PilotLight_Round_G_On_256c"; PictureOff "PilotLight_Round_G_Off_256c"
      ProcessValue <- "MS_IS2_SC_X1.4"
   TextField "Text field_35" at 536,146 size 114x20; Text 'MS_IS2_SC_X1.4'
   GraphicIOField "PlotLight_Round_G_35" at 664,168 size 24x24; PictureOn "PilotLight_Round_G_On_256c"; PictureOff "PilotLight_Round_G_Off_256c"
      ProcessValue <- "MS_IS2_SC_X1.5"
   TextField "Text field_36" at 536,170 size 114x20; Text 'MS_IS2_SC_X1.5'
   GraphicIOField "PlotLight_Round_G_36" at 664,192 size 24x24; PictureOn "PilotLight_Round_G_On_256c"; PictureOff "PilotLight_Round_G_Off_256c"
      ProcessValue <- "MS_IS2_SC_X1.6"
   TextField "Text field_37" at 536,194 size 114x20; Text 'MS_IS2_SC_X1.6'
   GraphicIOField "PlotLight_Round_G_37" at 664,216 size 24x24; PictureOn "PilotLight_Round_G_On_256c"; PictureOff "PilotLight_Round_G_Off_256c"
      ProcessValue <- "MS_IS2_SC_X1.7"
   TextField "Text field_38" at 536,218 size 114x20; Text 'MS_IS2_SC_X1.7'
   GraphicIOField "PlotLight_Round_G_38" at 488,240 size 24x24; PictureOff "PilotLight_Round_G_Off_256c"; PictureOn "PilotLight_Round_G_On_256c"
      ProcessValue <- "MS_OS_SC_X1.0"
   TextField "Text field_39" at 360,242 size 110x20; Text 'MS_OS_SC_X1.0'
   GraphicIOField "PlotLight_Round_G_39" at 488,264 size 24x24; PictureOn "PilotLight_Round_G_On_256c"; PictureOff "PilotLight_Round_G_Off_256c"
      ProcessValue <- "MS_OS_SC_X1.1"
   TextField "Text field_40" at 360,266 size 110x20; Text 'MS_OS_SC_X1.1'
   GraphicIOField "PlotLight_Round_G_40" at 488,288 size 24x24; PictureOn "PilotLight_Round_G_On_256c"; PictureOff "PilotLight_Round_G_Off_256c"
      ProcessValue <- "MS_OS_SC_X1.2"
   TextField "Text field_41" at 360,290 size 110x20; Text 'MS_OS_SC_X1.2'
   GraphicIOField "PlotLight_Round_G_41" at 488,312 size 24x24; PictureOff "PilotLight_Round_G_Off_256c"; PictureOn "PilotLight_Round_G_On_256c"
      ProcessValue <- "MS_OS_SC_X1.3"
   TextField "Text field_42" at 360,314 size 110x20; Text 'MS_OS_SC_X1.3'
   GraphicIOField "PlotLight_Round_G_42" at 488,336 size 24x24; PictureOff "PilotLight_Round_G_Off_256c"; PictureOn "PilotLight_Round_G_On_256c"
      ProcessValue <- "MS_OS_SC_X1.4"
   TextField "Text field_43" at 360,338 size 110x20; Text 'MS_OS_SC_X1.4'
   GraphicIOField "PlotLight_Round_G_43" at 488,360 size 24x24; PictureOff "PilotLight_Round_G_Off_256c"; PictureOn "PilotLight_Round_G_On_256c"
      ProcessValue <- "MS_OS_SC_X1.5"
   TextField "Text field_44" at 360,362 size 110x20; Text 'MS_OS_SC_X1.5'

screen "Manual.Destacker" 800x480, template "TemplateWithClockAndBackBtnForManual"
   on GenerateScreen: SetBit("Maintenance")
   on ClearScreen: ResetBit("Maintenance")
   TextField "Text field_14" at 496,54 size 179x20; Text 'Comanda 1 softstarter aer'
   TextField "Text field_15" at 496,134 size 190x20; Text 'Comanda cilindru vertical jos'
   TextField "Text field_16" at 496,174 size 193x20; Text 'Comanda cilindru vertical sus'
   TextField "Text field_17" at 496,214 size 155x20; Text 'Comanda furca retrasa'
   TextField "Text field_18" at 496,254 size 153x20; Text 'Comanda furca extinsa'
   Switch "Switch_1" at 696,128 size 64x32; CaptionText 'Switch'; TextOff 'OFF'; TextOn 'ON'
      ProcessValue <- "DS_Comanda cilindru vertical jos"
      on SwitchOn: SetBit("DS_Cilindru vertical jos")
      on SwitchOff: ResetBit("DS_Cilindru vertical jos")
   GraphicIOField "PlotLight_Round_G_2" at 160,48 size 24x24; PictureOn "PilotLight_Round_G_On_256c"; PictureOff "PilotLight_Round_G_Off_256c"
      ProcessValue <- "DB_PalletDispenser_PD2_De_Stacking_DB_PD1_MiddlePosition"
   TextField "Text field_3" at 16,50 size 126x20; Text 'PD1 MiddlePosition'
   Switch "Switch_2" at 696,48 size 64x32; CaptionText 'Switch'; TextOff 'OFF'; TextOn 'ON'
      ProcessValue <- "Comanda 1 softstarter aer destacker"
      on SwitchOn: SetBit("Comanda 1 softstarter aer destacker")
      on SwitchOff: ResetBit("Comanda 1 softstarter aer destacker")
   Switch "Switch_3" at 696,168 size 64x32; CaptionText 'Switch'; TextOff 'OFF'; TextOn 'ON'
      ProcessValue <- "DS_Comanda cilindru vertical sus"
      on SwitchOn: SetBit("DS_Cilindru vertical sus")
      on SwitchOff: ResetBit("DS_Cilindru vertical sus")
   Switch "Switch_4" at 696,208 size 64x32; CaptionText 'Switch'; TextOff 'OFF'; TextOn 'ON'
      ProcessValue <- "DS_Comanda furca retrasa"
      on SwitchOn: SetBit("DS_Comanda furca retrasa")
      on SwitchOff: ResetBit("DS_Comanda furca retrasa")
   Switch "Switch_5" at 696,248 size 64x32; CaptionText 'Switch'; TextOff 'OFF'; TextOn 'ON'
      ProcessValue <- "DS_Comanda furca extinsa"
      on SwitchOn: SetBit("DS_Comanda furca extinsa")
      on SwitchOff: ResetBit("DS_Comanda furca extinsa")
   TextField "Text field_21" at 496,94 size 179x20; Text 'Comanda 2 softstarter aer'
   Switch "Switch_8" at 696,88 size 64x32; CaptionText 'Switch'; TextOff 'OFF'; TextOn 'ON'
      ProcessValue <- "Comanda 2 softstarter aer destacker"
      on SwitchOn: SetBit("Comanda 2 softstarter aer destacker")
      on SwitchOff: ResetBit("Comanda 2 softstarter aer destacker")
   GraphicIOField "PlotLight_Round_G_1" at 160,72 size 24x24; PictureOff "PilotLight_Round_G_Off_256c"; PictureOn "PilotLight_Round_G_On_256c"
      ProcessValue <- "DB_PalletDispenser_PD2_De_Stacking_DB_PD1_Up"
   TextField "Text field_1" at 16,74 size 50x20; Text 'PD1 Up'
   GraphicIOField "PlotLight_Round_G_3" at 160,96 size 24x24; PictureOff "PilotLight_Round_G_Off_256c"; PictureOn "PilotLight_Round_G_On_256c"
      ProcessValue <- "DB_PalletDispenser_PD2_De_Stacking_DB_PD1_Down"
   TextField "Text field_2" at 16,98 size 70x20; Text 'PD1 Down'
   GraphicIOField "PlotLight_Round_G_4" at 160,120 size 24x24; PictureOff "PilotLight_Round_G_Off_256c"; PictureOn "PilotLight_Round_G_On_256c"
      ProcessValue <- "DB_PalletDispenser_PD2_De_Stacking_DB_PD1_Forks_In"
   TextField "Text field_4" at 16,122 size 85x20; Text 'PD1 Forks In'
   GraphicIOField "PlotLight_Round_G_5" at 160,144 size 24x24; PictureOn "PilotLight_Round_G_On_256c"; PictureOff "PilotLight_Round_G_Off_256c"
      ProcessValue <- "DB_PalletDispenser_PD2_De_Stacking_DB_PD1_Forks_Out"
   TextField "Text field_5" at 16,146 size 95x20; Text 'PD1 Forks Out'
   GraphicIOField "PlotLight_Round_G_7" at 160,167 size 24x24; PictureOff "PilotLight_Round_G_Off_256c"; PictureOn "PilotLight_Round_G_On_256c"
      ProcessValue <- "DB_PalletDispenser_PD2_De_Stacking_DB_Alarm_Active"
   TextField "Text field_7" at 16,169 size 89x20; Text 'Alarm Active'
   GraphicIOField "PlotLight_Round_G_8" at 416,48 size 24x24; PictureOn "PilotLight_Round_G_On_256c"; PictureOff "PilotLight_Round_G_Off_256c"
      ProcessValue <- "DS_Cilindru extins"
   TextField "Text field_8" at 240,50 size 120x20; Text 'DS_Cilindru extins'
   GraphicIOField "PlotLight_Round_G_9" at 416,72 size 24x24; PictureOn "PilotLight_Round_G_On_256c"; PictureOff "PilotLight_Round_G_Off_256c"
      ProcessValue <- "DS_Cilindru retras"
   TextField "Text field_9" at 240,74 size 122x20; Text 'DS_Cilindru retras'
   GraphicIOField "PlotLight_Round_G_10" at 416,96 size 24x24; PictureOff "PilotLight_Round_G_Off_256c"; PictureOn "PilotLight_Round_G_On_256c"
      ProcessValue <- "DS_Cilindru vertical jos"
   TextField "Text field_10" at 240,98 size 153x20; Text 'DS_Cilindru vertical jos'
   GraphicIOField "PlotLight_Round_G_11" at 416,120 size 24x24; PictureOff "PilotLight_Round_G_Off_256c"; PictureOn "PilotLight_Round_G_On_256c"
      ProcessValue <- "DS_Cilindru vertical mijloc"
   TextField "Text field_11" at 240,122 size 170x20; Text 'DS_Cilindru vertical mijloc'
   GraphicIOField "PlotLight_Round_G_12" at 416,144 size 24x24; PictureOff "PilotLight_Round_G_Off_256c"; PictureOn "PilotLight_Round_G_On_256c"
      ProcessValue <- "DS_Cilindru vertical sus"
   TextField "Text field_12" at 240,146 size 156x20; Text 'DS_Cilindru vertical sus'
   GraphicIOField "PlotLight_Round_G_13" at 416,168 size 24x24; PictureOn "PilotLight_Round_G_On_256c"; PictureOff "PilotLight_Round_G_Off_256c"
      ProcessValue <- "DS_Lungime 1"
   TextField "Text field_13" at 240,170 size 95x20; Text 'DS_Lungime 1'
   GraphicIOField "PlotLight_Round_G_14" at 416,192 size 24x24; PictureOn "PilotLight_Round_G_On_256c"; PictureOff "PilotLight_Round_G_Off_256c"
      ProcessValue <- "DS_Lungime 2"
   TextField "Text field_19" at 240,194 size 95x20; Text 'DS_Lungime 2'
   GraphicIOField "PlotLight_Round_G_15" at 416,216 size 24x24; PictureOff "PilotLight_Round_G_Off_256c"; PictureOn "PilotLight_Round_G_On_256c"
      ProcessValue <- "DS_Lungime 3"
   TextField "Text field_20" at 240,218 size 95x20; Text 'DS_Lungime 3'
   GraphicIOField "PlotLight_Round_G_29" at 416,240 size 24x24; PictureOn "PilotLight_Round_G_On_256c"; PictureOff "PilotLight_Round_G_Off_256c"
      ProcessValue <- "Senzor 1 proximitate softstarter aer destacker"
   TextField "Text field_30" at 96,242 size 312x20; Text 'Senzor 1 proximitate softstarter aer destacker'
   TextField "Text field_34" at 96,266 size 312x20; Text 'Senzor 2 proximitate softstarter aer destacker'